// TIA Portal project "New_V16_PID_Project_V5.5" (V16)

(* hardware
DEVICE "S7-1200 station_1"  S7-1200 Station
   slot 0: "Rack_0"  S7-1200 Rack  Rack  V1.0
   slot 1: "PLC_1"  CPU 1214C AC/DC/Rly  6ES7 214-1BG40-0XB0  V4.3
   slot 2: "AI 4xRTD_1"  SM 1231 AI4 x RTD  6ES7 231-5PD32-0XB0  V2.0
DEVICE "HMI_1"  TP1200 Comfort
   slot 0: "HMI_1"  TP1200 Comfort  6AV2 124-0MC01-0AX0  14.0.1.0
   slot 1: "HMI_RT_1"  TP1200 Comfort  6AV2 124-0MC01-0AX0  14.0.1.0
   slot 5: "HMI_1.IE_CP_1"  PROFINET Interface  14.0.1.0
      slot 1: "PROFINET Interface_1"  PROFINET Interface
         slot 1: "Port_1"  Port
         slot 2: "Port_2"  Port
   slot 7: "HMI_1.MPI/DP_CP_1"  MPI/DP Interface  14.0.1.0
*)

// ===== PLC "PLC_1"  CPU 1214C AC/DC/Rly =====

VAR_GLOBAL   // PLC tag table "Default tag table"
   "Start" AT %M0.0 : Bool;
   "Fan" AT %Q0.0 : Bool;
   "Fan Out Delay" AT %MD2 : Time;
   "Element Start" AT %M0.1 : Bool;
   "Element" AT %Q0.2 : Bool;
   "Element Time Delay" AT %MD6 : Time;
   "Start Up" AT %M0.2 : Bool;
   "Start Up Delay" AT %MD10 : Time;
   "Auger" AT %Q0.1 : Bool;
   "RTD" AT %IW96 : Word;
   "RTD 2" AT %IW98 : Word;
   "Setpoint" AT %MW20 : Word;
   "RTD Real" AT %MD14 : Real;
   "RTD 2 Real" AT %MD22 : Real;
   "Corrected RTD Temp" AT %MD26 : Real;
   "Corrected RTD 2 Temp" AT %MD30 : Real;
   "Auger PID" AT %M0.3 : Bool;
   "Corrected Setpoint" AT %MD34 : Real;
   "Auger Start Up" AT %M0.4 : Bool;
   "Auger Duty Cycle Start" AT %M0.5 : Bool;
   "Auger Duty Cycle" AT %M0.6 : Bool;
   "Auger Duty Cycle Output" AT %M0.7 : Bool;
   "Test Output" AT %M1.0 : Bool;
   "Set Reset" AT %M1.1 : Bool;
   "Error Ack" AT %M1.2 : Bool;
   "Error Ack Button" AT %M1.3 : Bool;
END_VAR

// folder: System blocks/Program resources

DATA_BLOCK "IEC_Timer_0_DB"   // DB1
{ S7_Optimized_Access := 'TRUE' }
AUTHOR : Simatic
FAMILY : IEC
NAME : IEC_TMR
VERSION : 1.0
// stored: InstanceOfName IEC_TIMER
"IEC_TIMER"
BEGIN
END_DATA_BLOCK

DATA_BLOCK "IEC_Timer_0_DB_1"   // DB3
{ S7_Optimized_Access := 'TRUE' }
AUTHOR : Simatic
FAMILY : IEC
NAME : IEC_TMR
VERSION : 1.0
// stored: InstanceOfName IEC_TIMER
"IEC_TIMER"
BEGIN
END_DATA_BLOCK

DATA_BLOCK "IEC_Timer_0_DB_2"   // DB5
{ S7_Optimized_Access := 'TRUE' }
AUTHOR : Simatic
FAMILY : IEC
NAME : IEC_TMR
VERSION : 1.0
// stored: InstanceOfName IEC_TIMER
"IEC_TIMER"
BEGIN
END_DATA_BLOCK

DATA_BLOCK "IEC_Timer_0_DB_3"   // DB9
{ S7_Optimized_Access := 'TRUE' }
AUTHOR : Simatic
FAMILY : IEC
NAME : IEC_TMR
VERSION : 1.0
// stored: InstanceOfName IEC_TIMER
"IEC_TIMER"
BEGIN
END_DATA_BLOCK

DATA_BLOCK "IEC_Timer_0_DB_4"   // DB10
{ S7_Optimized_Access := 'TRUE' }
AUTHOR : Simatic
FAMILY : IEC
NAME : IEC_TMR
VERSION : 1.0
// stored: InstanceOfName IEC_TIMER
"IEC_TIMER"
BEGIN
END_DATA_BLOCK

// folder: (top level)

ORGANIZATION_BLOCK "Main"   // OB1, LAD, ProgramCycle
TITLE = "Main Program Sweep (Cycle)"
{ S7_Optimized_Access := 'TRUE' }
VERSION : 0.1
   VAR_INPUT
      Initial_Call : Bool;   // Initial call of this OB
      Remanence : Bool;   // =True, if remanent data are available
   END_VAR
BEGIN

REGION Network 1
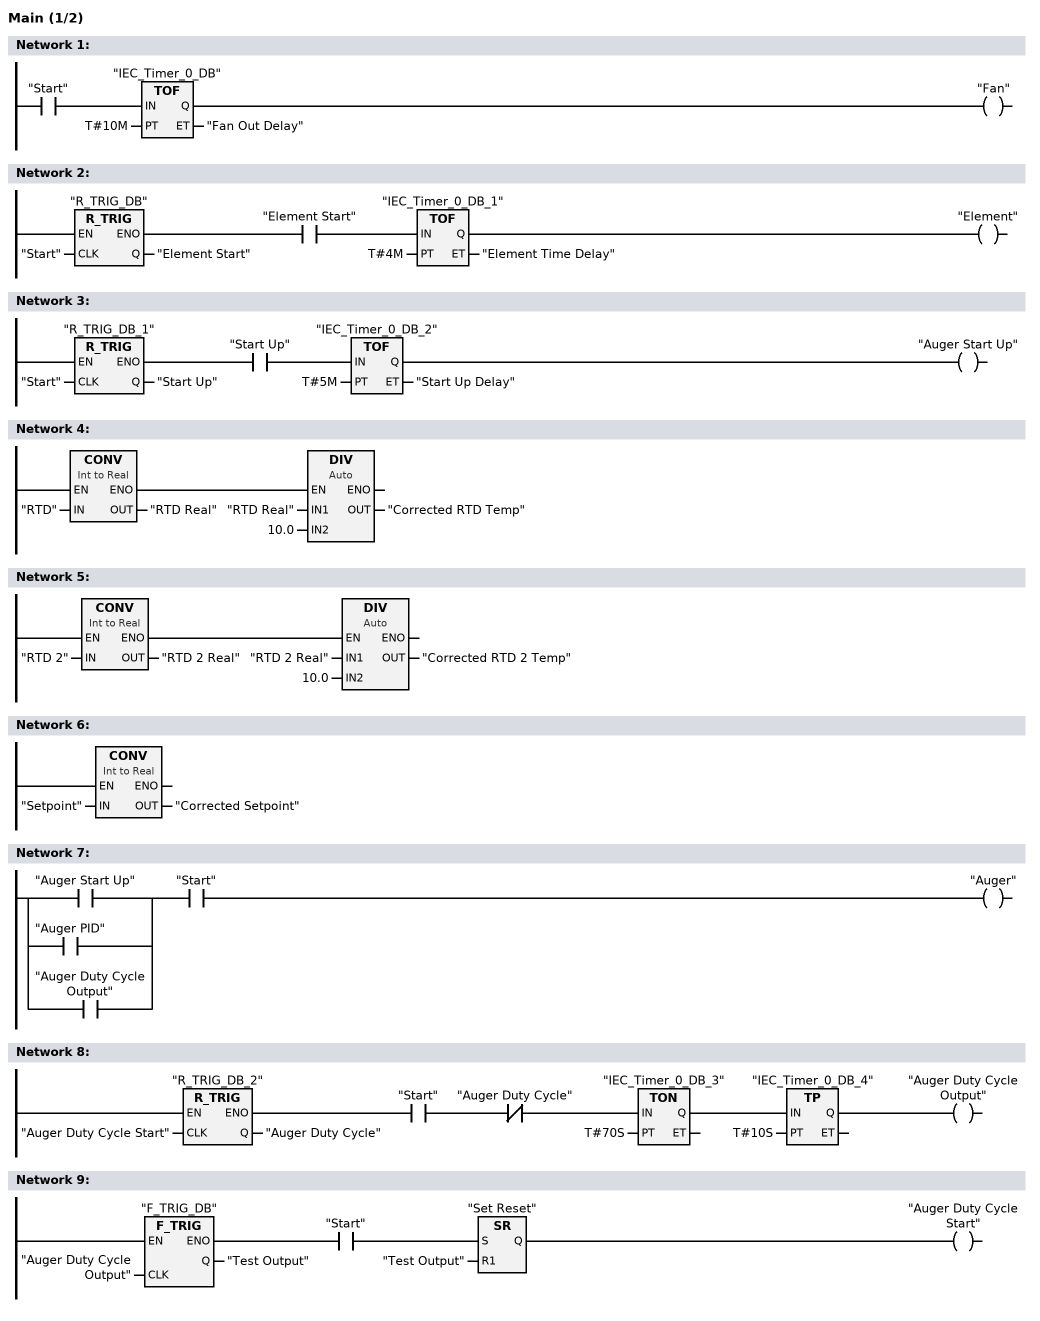
   "IEC_Timer_0_DB".TOF(IN := "Start", PT := T#10M, ET => "Fan Out Delay");
   "Fan" := "IEC_Timer_0_DB".Q;
END_REGION

REGION Network 2
   // ENO of a box is taken as its EN; it also drops when the box reports an error
   "R_TRIG_DB"(CLK := "Start", Q => "Element Start");   // R_TRIG
   "IEC_Timer_0_DB_1".TOF(IN := "Element Start", PT := T#4M, ET => "Element Time Delay");
   "Element" := "IEC_Timer_0_DB_1".Q;
END_REGION

REGION Network 3
   // ENO of a box is taken as its EN; it also drops when the box reports an error
   "R_TRIG_DB_1"(CLK := "Start", Q => "Start Up");   // R_TRIG
   "IEC_Timer_0_DB_2".TOF(IN := "Start Up", PT := T#5M, ET => "Start Up Delay");
   "Auger Start Up" := "IEC_Timer_0_DB_2".Q;
END_REGION

REGION Network 4
   RUNG wire#powerrail
      { S7_Templates := "[SrcType := Int, DestType := Real]" } Convert(in := "RTD", out => "RTD Real")
      Div(in1 := "RTD Real", in2 := 10.0, out => "Corrected RTD Temp")
   END_RUNG
   // the same network as SCL:
   "RTD Real" := INT_TO_REAL("RTD");
   "Corrected RTD Temp" := "RTD Real" / 10.0;
END_REGION

REGION Network 5
   RUNG wire#powerrail
      { S7_Templates := "[SrcType := Int, DestType := Real]" } Convert(in := "RTD 2", out => "RTD 2 Real")
      Div(in1 := "RTD 2 Real", in2 := 10.0, out => "Corrected RTD 2 Temp")
   END_RUNG
   // the same network as SCL:
   "RTD 2 Real" := INT_TO_REAL("RTD 2");
   "Corrected RTD 2 Temp" := "RTD 2 Real" / 10.0;
END_REGION

REGION Network 6
   RUNG wire#powerrail
      { S7_Templates := "[SrcType := Int, DestType := Real]" } Convert(in := "Setpoint", out => "Corrected Setpoint")
   END_RUNG
   // the same network as SCL:
   "Corrected Setpoint" := INT_TO_REAL("Setpoint");
END_REGION

REGION Network 7
   RUNG wire#powerrail
      Contact( "Auger Start Up" )
      wire#w1
      Contact( "Start" )
      Coil( "Auger" )
   END_RUNG
   RUNG wire#powerrail
      Contact( "Auger PID" )
   END_RUNG wire#w1
   RUNG wire#powerrail
      Contact( "Auger Duty Cycle Output" )
   END_RUNG wire#w1
   // the same network as SCL:
   "Auger" := ("Auger Start Up" OR "Auger PID" OR "Auger Duty Cycle Output") AND "Start";
END_REGION

REGION Network 8
   // ENO of a box is taken as its EN; it also drops when the box reports an error
   "R_TRIG_DB_2"(CLK := "Auger Duty Cycle Start", Q => "Auger Duty Cycle");   // R_TRIG
   "IEC_Timer_0_DB_3".TON(IN := "Start" AND NOT "Auger Duty Cycle", PT := T#70S);
   "IEC_Timer_0_DB_4".TP(IN := "IEC_Timer_0_DB_3".Q, PT := T#10S);
   "Auger Duty Cycle Output" := "IEC_Timer_0_DB_4".Q;
END_REGION

REGION Network 9
   // ENO of a box is taken as its EN; it also drops when the box reports an error
   "F_TRIG_DB"(CLK := "Auger Duty Cycle Output", Q => "Test Output");   // F_TRIG
   IF "Start" THEN
       "Set Reset" := TRUE;   // SR flip-flop
   END_IF;
   IF "Test Output" THEN "Set Reset" := FALSE; END_IF;
   "Auger Duty Cycle Start" := "Set Reset";
END_REGION

REGION Network 10
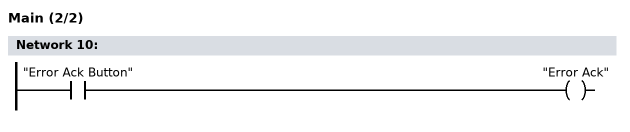
   RUNG wire#powerrail
      Contact( "Error Ack Button" )
      Coil( "Error Ack" )
   END_RUNG
   // the same network as SCL:
   "Error Ack" := "Error Ack Button";
END_REGION
END_ORGANIZATION_BLOCK

ORGANIZATION_BLOCK "Cyclic interrupt"   // OB30, LAD, CyclicInterrupt
{ S7_Optimized_Access := 'TRUE' }
VERSION : 0.1
   VAR_INPUT
      Initial_Call : Bool;   // Initial call of this OB
      Event_Count : Int;   // Events discarded
   END_VAR
BEGIN

REGION Network 1
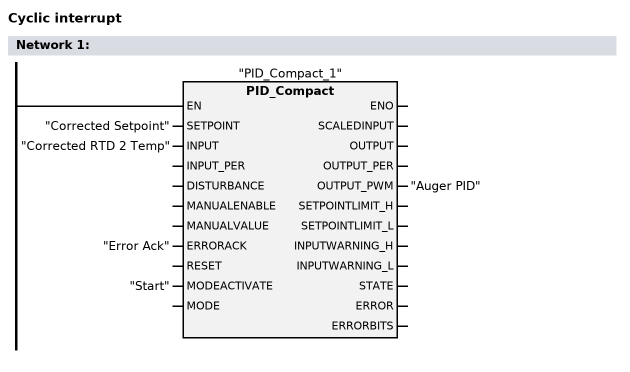
   "PID_Compact_1"(Setpoint := "Corrected Setpoint",   // PID_Compact
                   Input := "Corrected RTD 2 Temp",
                   ErrorAck := "Error Ack",
                   ModeActivate := "Start",
                   Output_PWM => "Auger PID");
END_REGION
END_ORGANIZATION_BLOCK

(* ===== HMI "HMI_RT_1" =====
system functions are stored by id; their names below are inferred from use
connection "HMI_Connection_1": ETHERNET, S7_1200_OMS

HMI tags "Default tag table"
   "Tag_ScreenNumber" : UInt, internal
   "Start" : Bool = PLC Start AT %M0.0, 1 s
   "Setpoint" : Word = PLC Setpoint AT %MW20, 1 s
   "Corrected RTD 2 Temp" : Real = PLC "Corrected RTD 2 Temp" AT %MD30, 1 s
   "Error Ack Button" : Bool = PLC "Error Ack Button" AT %M1.3, 1 s

screen "Root screen" 1280x740, template "Template_1"
   on GenerateScreen: SetTag("Tag_ScreenNumber", 1)
   Switch "Switch_1" at 118,452 size 204x144; CaptionText 'Smoker Switch'; TextOff 'OFF'; TextOn 'ON'
      ProcessValue <- "Start"
   Button "Button_1" at 104,54 size 222x72; TextOff 'RUN'
      on Click: function_f249594b("HMI_Connection_1", 8)
   Button "Button_2" at 104,161 size 224x74; TextOff 'STOP'
      on Click: function_f249594b("HMI_Connection_1", 4)
   Gauge "Gauge_1" at 868,178 size 304x304; CaptionText 'RTD Temp'; UnitText 'Fahrenheit'
      ProcessValue <- "Corrected RTD 2 Temp"
   Button "Button_3" at 105,275 size 223x72; TextOff 'Error Ack'
      on Press: function_b14e0dd5("Error Ack Button", 0)
   Slider "Slider_1" at 496,22 size 214x644; Caption 'Set Point Temp'
      ProcessValue <- "Setpoint"

Template "Template_1" 1280x740
   Button "Exit" at 1200,679 size 78x59; TextOff 'Exit'; PictureOff "ExitRuntime_TP1200_Comfort_TR"; PictureOn "ExitRuntime_TP1200_Comfort_TR"
      on Release: StopRuntime(0)
   Button "Template_Button" at 1120,679 size 78x59; TextOff 'Text'
   Button "Template_Button_1" at 1040,679 size 78x59; TextOff 'Text'
   Button "Template_Button_2" at 960,679 size 78x59; TextOff 'Text'
   Button "Template_Button_3" at 880,679 size 78x59; TextOff 'Text'
   Button "Template_Button_4" at 800,679 size 78x59; TextOff 'Text'
   Button "Template_Button_5" at 720,679 size 78x59; TextOff 'Text'
   Button "Template_Button_6" at 640,679 size 78x59; TextOff 'Text'
   Button "Template_Button_7" at 561,679 size 78x59; TextOff 'Text'
   Button "Template_Button_8" at 481,679 size 78x59; TextOff 'Text'
   Button "Template_Button_9" at 401,679 size 78x59; TextOff 'Text'
   Button "Template_Button_10" at 321,679 size 78x59; TextOff 'Text'
   Button "Template_Button_11" at 241,679 size 78x59; TextOff 'Text'
   Button "Template_Button_12" at 161,679 size 78x59; TextOff 'Text'
   Button "Alarms" at 81,679 size 78x59; TextOff 'Alarms'; PictureOff "AlarmDisplay_TP1200_Comfort_TR"; PictureOn "AlarmDisplay_TP1200_Comfort_TR"
      on Release: function_ef3f5d25("Alarm window_Unacknowledged", -1)
   Button "Start screen" at 1,679 size 78x59; TextOff 'Start screen'; PictureOff "NavigateHome_TP1200_Comfort_TR"; PictureOn "NavigateHome_TP1200_Comfort_TR"
      on Release: ActivateScreen("Root screen", 0)
*)